(* Logix 5000 project; controller FV vendor 1 type 14 code 217 rev 31.11; software revision 31.00; part 4 of 63 *)

        [1]   // FV12,TEMPERATURE BREAKPOINT A. TIME 1/10 HOURS(ALWAYS=0)
        [15].5   // FV12,Profile Control Flags : This is a conditioning profile
        [29].1   // FV12,Current vessel deferred chilling enabled flag
        [3]   // FV12,TEMPERATURE BREAKPOINT B. TIME 1/10 HOURS(ALWAYS=0)
        [5]   // FV12,TEMPERATURE BREAKPOINT C. TIME 1/10 HOURS(ALWAYS=0)
        [7]   // FV12,TEMPERATURE BREAKPOINT D. TIME 1/10 HOURS(ALWAYS=0)
        [9]   // FV12,TEMPERATURE BREAKPOINT E. TIME 1/10 HOURS(ALWAYS=0)
        [15].9   // FV12,Current vessel deferred chilling manual override
   FV_N123 : INT[50] := ([0] := 13, [2] := 170, [3] := 100, [4] := 190, [5] := 245, [6] := 190, [7] := 275, [8] := 160, [9] := 480, [10] := 160, [11] := 580, [12] := 60, [13] := 32767, [14] := 60, [15] := 64, [17] := -32767, [18] := -32767, [19] := 1680, [22] := 487, [23] := 3, [24] := 5, [25] := 153, [26] := 153, [27] := 487, [30] := 1);   // FV13, CURRENT FV DATA
        [15].2   // FV13,PLC TO FOLLOW RAMP Breakpoints A to B
        [15]   // FV13,FLAGS-PROFILE CONTROL
        [41]   // FV13,Cone ACTUAL TEMPERATURE -DEGREES 'C'*10
        [28]   // FV13,CURRENT VOLUME HL*10
        [15].3   // FV13,PLC TO USE CONE COOLING JACKET
        [24]   // FV13,Phase0=No control 1to6 =Fermenting 8 =Pitching Hold 10 =Maturation 11to16=Conditioning
        [26]   // FV13,Calculated Setpoint 1/10 degrees C
        [30].1   // FV13,Cone Cooling Valve to open
        [30].0   // FV13,Jacket Cooling Valve to open
        [19]   // FV13,Current FV max. fermentation time
        [25]   // FV13,Jacket ACTUAL TEMPERATURE -DEGREES 'C'*10
        [20]   // FV13,Current FV warm conditioning time
        [29]   // FV13,FLAGS - PLC CONTROL
        [10]   // FV13,TEMPERATURE SETPOINT E. 1/10 DEGREE 'C'
        [12]   // FV13,TEMPERATURE SETPOINT F. 1/10 DEGREE 'C'
        [14]   // FV13,TEMPERATURE SETPOINT G. 1/10 DEGREE 'C'
        [30].3   // FV13,Current vessel deferred chilling active
        [0]   // FV13,FV SYSTEM WORKING BUFFER VESSEL NUMBER
        [2]   // FV13,TEMPERATURE SETPOINT A. 1/10 DEGREE 'C'
        [30].4   // FV13,Current vessel final temp.reached
        [4]   // FV13,TEMPERATURE SETPOINT B. 1/10 DEGREE 'C'
        [6]   // FV13,TEMPERATURE SETPOINT C. 1/10 DEGREE 'C'
        [8]   // FV13,TEMPERATURE SETPOINT D. 1/10 DEGREE 'C'
        [22]   // FV13,Current FV total residence time
        [29].0   // FV13,PC TO SAVE TEMPERATURE DATA
        [11]   // FV13,TEMPERATURE BREAKPOINT F. TIME 1/10 HOURS(ALWAYS=0)
        [13]   // FV13,TEMPERATURE BREAKPOINT G. TIME 1/10 HOURS(ALWAYS=0)
        [30].5   // FV13,Current vessel deferred chilling temp.high flag
        [16].1   // FV13,Profile control flag Hold at B.P B
        [16].2   // FV13,Profile control flag Hold at B.P C
        [16].3   // FV13,Profile control flag Hold at B.P D
        [16].4   // FV13,Profile control flag Hold at B.P E
        [16].5   // FV13,Profile control flag Hold at B.P F
        [16].6   // FV13,Profile control flag Hold at B.P G
        [15].4   // FV13,Profile Control Flags : This is a maturation profile
        [27]   // FV13,CURRENT ELAPSED HOURS *10
        [40]   // FV13,FV Routing Status 9=Dirty
        [15].5   // FV13,Profile Control Flags : This is a conditioning profile
        [36]   // FV13,Current vessel time to deferred chlling start (hrs.x10)
        [1]   // FV13,TEMPERATURE BREAKPOINT A. TIME 1/10 HOURS(ALWAYS=0)
        [29].1   // FV13,Current vessel deferred chilling enabled flag
        [3]   // FV13,TEMPERATURE BREAKPOINT B. TIME 1/10 HOURS(ALWAYS=0)
        [5]   // FV13,TEMPERATURE BREAKPOINT C. TIME 1/10 HOURS(ALWAYS=0)
        [7]   // FV13,TEMPERATURE BREAKPOINT D. TIME 1/10 HOURS(ALWAYS=0)
        [9]   // FV13,TEMPERATURE BREAKPOINT E. TIME 1/10 HOURS(ALWAYS=0)
        [15].9   // FV13,Current vessel deferred chilling manual override
   FV_N124 : INT[50] := ([0] := 14, [2] := 170, [3] := 100, [4] := 190, [5] := 258, [6] := 190, [7] := 290, [8] := 160, [9] := 505, [10] := 160, [11] := 605, [12] := 60, [13] := 32767, [14] := 60, [15] := 64, [17] := -32767, [18] := -32767, [19] := 1680, [20] := 8, [22] := 1688, [23] := 3, [24] := 6, [25] := 62, [26] := 60, [27] := 1688, [29] := 2, [30] := 24);   // FV14, CURRENT FV DATA
        [15]   // FV14,FLAGS-PROFILE CONTROL
        [15].2   // FV14,PLC TO FOLLOW RAMP Breakpoints A to B
        [41]   // FV14,Cone ACTUAL TEMPERATURE -DEGREES 'C'*10
        [28]   // FV14,CURRENT VOLUME HL*10
        [30].1   // FV14,Cone Cooling Valve to open
        [15].3   // FV14,PLC TO USE CONE COOLING JACKET
        [24]   // FV14,Phase0=No control 1to6 =Fermenting 8 =Pitching Hold 10 =Maturation 11to16=Conditioning
        [25]   // FV14,Jacket ACTUAL TEMPERATURE -DEGREES 'C'*10
        [26]   // FV14,Calculated Setpoint 1/10 degrees C
        [30].0   // FV14,Jacket Cooling Valve to open
        [19]   // FV14,Current FV max. fermentation time
        [20]   // FV14,Current FV warm conditioning time
        [29]   // FV14,FLAGS - PLC CONTROL
        [0]   // FV14,FV SYSTEM WORKING BUFFER VESSEL NUMBER
        [10]   // FV14,TEMPERATURE SETPOINT E. 1/10 DEGREE 'C'
        [12]   // FV14,TEMPERATURE SETPOINT F. 1/10 DEGREE 'C'
        [2]   // FV14,TEMPERATURE SETPOINT A. 1/10 DEGREE 'C'
        [14]   // FV14,TEMPERATURE SETPOINT G. 1/10 DEGREE 'C'
        [30].3   // FV14,Current vessel deferred chilling active
        [30].4   // FV14,Current vessel final temp.reached
        [4]   // FV14,TEMPERATURE SETPOINT B. 1/10 DEGREE 'C'
        [6]   // FV14,TEMPERATURE SETPOINT C. 1/10 DEGREE 'C'
        [8]   // FV14,TEMPERATURE SETPOINT D. 1/10 DEGREE 'C'
        [22]   // FV14,Current FV total residence time
        [29].0   // FV14,PC TO SAVE TEMPERATURE DATA
        [11]   // FV14,TEMPERATURE BREAKPOINT F. TIME 1/10 HOURS(ALWAYS=0)
        [13]   // FV14,TEMPERATURE BREAKPOINT G. TIME 1/10 HOURS(ALWAYS=0)
        [30].5   // FV14,Current vessel deferred chilling temp.high flag
        [16].1   // FV14,Profile control flag Hold at B.P B
        [16].2   // FV14,Profile control flag Hold at B.P C
        [16].3   // FV14,Profile control flag Hold at B.P D
        [16].4   // FV14,Profile control flag Hold at B.P E
        [16].5   // FV14,Profile control flag Hold at B.P F
        [16].6   // FV14,Profile control flag Hold at B.P G
        [27]   // FV14,CURRENT ELAPSED HOURS *10
        [40]   // FV14,FV Routing Status 9=Dirty
        [15].4   // FV14,Profile Control Flags : This is a maturation profile
        [15].5   // FV14,Profile Control Flags : This is a conditioning profile
        [36]   // FV14,Current vessel time to deferred chlling start (hrs.x10)
        [15].9   // FV14,Current vessel deferred chilling manual override
        [1]   // FV14,TEMPERATURE BREAKPOINT A. TIME 1/10 HOURS(ALWAYS=0)
        [29].1   // FV14,Current vessel deferred chilling enabled flag
        [3]   // FV14,TEMPERATURE BREAKPOINT B. TIME 1/10 HOURS(ALWAYS=0)
        [5]   // FV14,TEMPERATURE BREAKPOINT C. TIME 1/10 HOURS(ALWAYS=0)
        [7]   // FV14,TEMPERATURE BREAKPOINT D. TIME 1/10 HOURS(ALWAYS=0)
        [9]   // FV14,TEMPERATURE BREAKPOINT E. TIME 1/10 HOURS(ALWAYS=0)
   FV_N125 : INT[50] := ([0] := 15, [2] := 170, [3] := 100, [4] := 190, [5] := 270, [6] := 190, [7] := 300, [8] := 160, [9] := 530, [10] := 160, [11] := 630, [12] := 60, [13] := 32767, [14] := 60, [15] := 64, [16] := 20, [17] := -32767, [18] := -32767, [19] := 1680, [22] := 8, [23] := 1, [24] := 1, [25] := 174, [26] := 190, [27] := 8);   // FV15, CURRENT FV DATA
        [15]   // FV15,FLAGS-PROFILE CONTROL
        [15].2   // FV15,PLC TO FOLLOW RAMP Breakpoints A to B
        [41]   // FV15,Cone ACTUAL TEMPERATURE -DEGREES 'C'*10
        [28]   // FV15,CURRENT VOLUME HL*10
        [30].0   // FV15,Jacket Cooling Valve to open
        [30].1   // FV15,Cone Cooling Valve to open
        [15].3   // FV15,PLC TO USE CONE COOLING JACKET
        [24]   // FV15,Phase0=No control 1to6 =Fermenting 8 =Pitching Hold 10 =Maturation 11to16=Conditioning
        [25]   // FV15,Jacket ACTUAL TEMPERATURE -DEGREES 'C'*10
        [26]   // FV15,Calculated Setpoint 1/10 degrees C
        [19]   // FV15,Current FV max. fermentation time
        [20]   // FV15,Current FV warm conditioning time
        [29]   // FV15,FLAGS - PLC CONTROL
        [10]   // FV15,TEMPERATURE SETPOINT E. 1/10 DEGREE 'C'
        [0]   // FV15,FV SYSTEM WORKING BUFFER VESSEL NUMBER
        [2]   // FV15,TEMPERATURE SETPOINT A. 1/10 DEGREE 'C'
        [12]   // FV15,TEMPERATURE SETPOINT F. 1/10 DEGREE 'C'
        [30].4   // FV15,Current vessel final temp.reached
        [14]   // FV15,TEMPERATURE SETPOINT G. 1/10 DEGREE 'C'
        [4]   // FV15,TEMPERATURE SETPOINT B. 1/10 DEGREE 'C'
        [6]   // FV15,TEMPERATURE SETPOINT C. 1/10 DEGREE 'C'
        [8]   // FV15,TEMPERATURE SETPOINT D. 1/10 DEGREE 'C'
        [30].3   // FV15,Current vessel deferred chilling active
        [22]   // FV15,Current FV total residence time
        [29].0   // FV15,PC TO SAVE TEMPERATURE DATA
        [11]   // FV15,TEMPERATURE BREAKPOINT F. TIME 1/10 HOURS(ALWAYS=0)
        [13]   // FV15,TEMPERATURE BREAKPOINT G. TIME 1/10 HOURS(ALWAYS=0)
        [30].5   // FV15,Current vessel deferred chilling temp.high flag
        [16].1   // FV15,Profile control flag Hold at B.P B
        [16].2   // FV15,Profile control flag Hold at B.P C
        [16].3   // FV15,Profile control flag Hold at B.P D
        [16].4   // FV15,Profile control flag Hold at B.P E
        [16].5   // FV15,Profile control flag Hold at B.P F
        [16].6   // FV15,Profile control flag Hold at B.P G
        [15].4   // FV15,Profile Control Flags : This is a maturation profile
        [15].5   // FV15,Profile Control Flags : This is a conditioning profile
        [27]   // FV15,CURRENT ELAPSED HOURS *10
        [40]   // FV15,FV Routing Status 9=Dirty
        [36]   // FV15,Current vessel time to deferred chlling start (hrs.x10)
        [15].9   // FV15,Current vessel deferred chilling manual override
        [1]   // FV15,TEMPERATURE BREAKPOINT A. TIME 1/10 HOURS(ALWAYS=0)
        [29].1   // FV15,Current vessel deferred chilling enabled flag
        [3]   // FV15,TEMPERATURE BREAKPOINT B. TIME 1/10 HOURS(ALWAYS=0)
        [5]   // FV15,TEMPERATURE BREAKPOINT C. TIME 1/10 HOURS(ALWAYS=0)
        [7]   // FV15,TEMPERATURE BREAKPOINT D. TIME 1/10 HOURS(ALWAYS=0)
        [9]   // FV15,TEMPERATURE BREAKPOINT E. TIME 1/10 HOURS(ALWAYS=0)
   FV_N126 : INT[50] := ([0] := 16, [1] := -32767, [2] := -32767, [3] := -32767, [4] := -32767, [5] := -32767, [6] := -32767, [7] := -32767, [8] := -32767, [9] := -32767, [10] := -32767, [11] := -32767, [12] := -32767, [13] := -32767, [14] := -32767, [15] := -32767, [16] := -32767, [17] := -32767, [18] := -32767, [19] := -32767, [20] := -32767, [21] := -32767, [22] := -32767, [23] := 2, [25] := 201, [30] := 32);   // FV16, CURRENT FV DATA
        [15]   // FV16,FLAGS-PROFILE CONTROL
        [15].2   // FV16,PLC TO FOLLOW RAMP Breakpoints A to B
        [41]   // FV16,Cone ACTUAL TEMPERATURE -DEGREES 'C'*10
        [28]   // FV16,CURRENT VOLUME HL*10
        [25]   // FV16,Jacket ACTUAL TEMPERATURE -DEGREES 'C'*10
        [15].3   // FV16,PLC TO USE CONE COOLING JACKET
        [30].0   // FV16,Jacket Cooling Valve to open
        [26]   // FV16,Calculated Setpoint 1/10 degrees C
        [30].1   // FV16,Cone Cooling Valve to open
        [24]   // FV16,Phase0=No control 1to6 =Fermenting 8 =Pitching Hold 10 =Maturation 11to16=Conditioning
        [19]   // FV16,Current FV max. fermentation time
        [20]   // FV16,Current FV warm conditioning time
        [29]   // FV16,FLAGS - PLC CONTROL
        [10]   // FV16,TEMPERATURE SETPOINT E. 1/10 DEGREE 'C'
        [12]   // FV16,TEMPERATURE SETPOINT F. 1/10 DEGREE 'C'
        [14]   // FV16,TEMPERATURE SETPOINT G. 1/10 DEGREE 'C'
        [0]   // FV16,FV SYSTEM WORKING BUFFER VESSEL NUMBER
        [2]   // FV16,TEMPERATURE SETPOINT A. 1/10 DEGREE 'C'
        [30].4   // FV16,Current vessel final temp.reached
        [4]   // FV16,TEMPERATURE SETPOINT B. 1/10 DEGREE 'C'
        [6]   // FV16,TEMPERATURE SETPOINT C. 1/10 DEGREE 'C'
        [8]   // FV16,TEMPERATURE SETPOINT D. 1/10 DEGREE 'C'
        [30].3   // FV16,Current vessel deferred chilling active
        [22]   // FV16,Current FV total residence time
        [29].0   // FV16,PC TO SAVE TEMPERATURE DATA
        [11]   // FV16,TEMPERATURE BREAKPOINT F. TIME 1/10 HOURS(ALWAYS=0)
        [13]   // FV16,TEMPERATURE BREAKPOINT G. TIME 1/10 HOURS(ALWAYS=0)
        [30].5   // FV16,Current vessel deferred chilling temp.high flag
        [36]   // FV16,Current vessel time to deferred chlling start (hrs.x10)
        [15].4   // FV16,Profile Control Flags : This is a maturation profile
        [15].5   // FV16,Profile Control Flags : This is a conditioning profile
        [16].1   // FV16,Profile control flag Hold at B.P B
        [16].2   // FV16,Profile control flag Hold at B.P C
        [16].3   // FV16,Profile control flag Hold at B.P D
        [16].4   // FV16,Profile control flag Hold at B.P E
        [16].5   // FV16,Profile control flag Hold at B.P F
        [16].6   // FV16,Profile control flag Hold at B.P G
        [27]   // FV16,CURRENT ELAPSED HOURS *10
        [40]   // FV16,FV Routing Status 9=Dirty
        [15].9   // FV16,Current vessel deferred chilling manual override
        [1]   // FV16,TEMPERATURE BREAKPOINT A. TIME 1/10 HOURS(ALWAYS=0)
        [29].1   // FV16,Current vessel deferred chilling enabled flag
        [3]   // FV16,TEMPERATURE BREAKPOINT B. TIME 1/10 HOURS(ALWAYS=0)
        [5]   // FV16,TEMPERATURE BREAKPOINT C. TIME 1/10 HOURS(ALWAYS=0)
        [7]   // FV16,TEMPERATURE BREAKPOINT D. TIME 1/10 HOURS(ALWAYS=0)
        [9]   // FV16,TEMPERATURE BREAKPOINT E. TIME 1/10 HOURS(ALWAYS=0)
   FV_N127 : INT[50] := ([0] := 17, [1] := -32767, [2] := -32767, [3] := -32767, [4] := -32767, [5] := -32767, [6] := -32767, [7] := -32767, [8] := -32767, [9] := -32767, [10] := -32767, [11] := -32767, [12] := -32767, [13] := -32767, [14] := -32767, [15] := -32767, [16] := -32767, [17] := -32767, [18] := -32767, [19] := -32767, [20] := -32767, [21] := -32767, [22] := -32767, [23] := 2, [25] := 203, [30] := 32);   // FV17, CURRENT FV DATA
        [15]   // FV17,FLAGS-PROFILE CONTROL
        [15].2   // FV17,PLC TO FOLLOW RAMP Breakpoints A to B
        [41]   // FV17,Cone ACTUAL TEMPERATURE -DEGREES 'C'*10
        [25]   // FV17,Jacket ACTUAL TEMPERATURE -DEGREES 'C'*10
        [28]   // FV17,CURRENT VOLUME HL*10
        [15].3   // FV17,PLC TO USE CONE COOLING JACKET
        [30].0   // FV17,Jacket Cooling Valve to open
        [26]   // FV17,Calculated Setpoint 1/10 degrees C
        [24]   // FV17,Phase0=No control 1to6 =Fermenting 8 =Pitching Hold 10 =Maturation 11to16=Conditioning
        [30].1   // FV17,Cone Cooling Valve to open
        [19]   // FV17,Current FV max. fermentation time
        [10]   // FV17,TEMPERATURE SETPOINT E. 1/10 DEGREE 'C'
        [20]   // FV17,Current FV warm conditioning time
        [12]   // FV17,TEMPERATURE SETPOINT F. 1/10 DEGREE 'C'
        [29]   // FV17,FLAGS - PLC CONTROL
        [14]   // FV17,TEMPERATURE SETPOINT G. 1/10 DEGREE 'C'
        [0]   // FV17,FV SYSTEM WORKING BUFFER VESSEL NUMBER
        [2]   // FV17,TEMPERATURE SETPOINT A. 1/10 DEGREE 'C'
        [30].4   // FV17,Current vessel final temp.reached
        [4]   // FV17,TEMPERATURE SETPOINT B. 1/10 DEGREE 'C'
        [6]   // FV17,TEMPERATURE SETPOINT C. 1/10 DEGREE 'C'
        [8]   // FV17,TEMPERATURE SETPOINT D. 1/10 DEGREE 'C'
        [30].3   // FV17,Current vessel deferred chilling active
        [22]   // FV17,Current FV total residence time
        [29].0   // FV17,PC TO SAVE TEMPERATURE DATA
        [36]   // FV17,Current vessel time to deferred chlling start (hrs.x10)
        [11]   // FV17,TEMPERATURE BREAKPOINT F. TIME 1/10 HOURS(ALWAYS=0)
        [13]   // FV17,TEMPERATURE BREAKPOINT G. TIME 1/10 HOURS(ALWAYS=0)
        [30].5   // FV17,Current vessel deferred chilling temp.high flag
        [15].4   // FV17,Profile Control Flags : This is a maturation profile
        [27]   // FV17,CURRENT ELAPSED HOURS *10
        [40]   // FV17,FV Routing Status 9=Dirty
        [16].1   // FV17,Profile control flag Hold at B.P B
        [15].5   // FV17,Profile Control Flags : This is a conditioning profile
        [16].2   // FV17,Profile control flag Hold at B.P C
        [16].3   // FV17,Profile control flag Hold at B.P D
        [16].4   // FV17,Profile control flag Hold at B.P E
        [16].5   // FV17,Profile control flag Hold at B.P F
        [16].6   // FV17,Profile control flag Hold at B.P G
        [15].9   // FV17,Current vessel deferred chilling manual override
        [1]   // FV17,TEMPERATURE BREAKPOINT A. TIME 1/10 HOURS(ALWAYS=0)
        [29].1   // FV17,Current vessel deferred chilling enabled flag
        [3]   // FV17,TEMPERATURE BREAKPOINT B. TIME 1/10 HOURS(ALWAYS=0)
        [5]   // FV17,TEMPERATURE BREAKPOINT C. TIME 1/10 HOURS(ALWAYS=0)
        [7]   // FV17,TEMPERATURE BREAKPOINT D. TIME 1/10 HOURS(ALWAYS=0)
        [9]   // FV17,TEMPERATURE BREAKPOINT E. TIME 1/10 HOURS(ALWAYS=0)
   FV_N128 : INT[50] := ([0] := 18, [1] := -32767, [2] := -32767, [3] := -32767, [4] := -32767, [5] := -32767, [6] := -32767, [7] := -32767, [8] := -32767, [9] := -32767, [10] := -32767, [11] := -32767, [12] := -32767, [13] := -32767, [14] := -32767, [15] := -32767, [16] := -32767, [17] := -32767, [18] := -32767, [19] := -32767, [20] := -32767, [21] := -32767, [22] := -32767, [23] := 2, [25] := 216, [30] := 32);   // FV18, CURRENT FV DATA
        [15]   // FV18,FLAGS-PROFILE CONTROL
        [15].2   // FV18,PLC TO FOLLOW RAMP Breakpoints A to B
        [25]   // FV18,Jacket ACTUAL TEMPERATURE -DEGREES 'C'*10
        [41]   // FV18,Cone ACTUAL TEMPERATURE -DEGREES 'C'*10
        [28]   // FV18,CURRENT VOLUME HL*10
        [15].3   // FV18,PLC TO USE CONE COOLING JACKET
        [26]   // FV18,Calculated Setpoint 1/10 degrees C
        [30].0   // FV18,Jacket Cooling Valve to open
        [30].1   // FV18,Cone Cooling Valve to open
        [24]   // FV18,Phase0=No control 1to6 =Fermenting 8 =Pitching Hold 10 =Maturation 11to16=Conditioning
        [19]   // FV18,Current FV max. fermentation time
        [20]   // FV18,Current FV warm conditioning time
        [10]   // FV18,TEMPERATURE SETPOINT E. 1/10 DEGREE 'C'
        [12]   // FV18,TEMPERATURE SETPOINT F. 1/10 DEGREE 'C'
        [14]   // FV18,TEMPERATURE SETPOINT G. 1/10 DEGREE 'C'
        [29]   // FV18,FLAGS - PLC CONTROL
        [0]   // FV18,FV SYSTEM WORKING BUFFER VESSEL NUMBER
        [2]   // FV18,TEMPERATURE SETPOINT A. 1/10 DEGREE 'C'
        [30].4   // FV18,Current vessel final temp.reached
        [4]   // FV18,TEMPERATURE SETPOINT B. 1/10 DEGREE 'C'
        [6]   // FV18,TEMPERATURE SETPOINT C. 1/10 DEGREE 'C'
        [8]   // FV18,TEMPERATURE SETPOINT D. 1/10 DEGREE 'C'
        [30].3   // FV18,Current vessel deferred chilling active
        [22]   // FV18,Current FV total residence time
        [29].0   // FV18,PC TO SAVE TEMPERATURE DATA
        [36]   // FV18,Current vessel time to deferred chlling start (hrs.x10)
        [15].4   // FV18,Profile Control Flags : This is a maturation profile
        [15].5   // FV18,Profile Control Flags : This is a conditioning profile
        [11]   // FV18,TEMPERATURE BREAKPOINT F. TIME 1/10 HOURS(ALWAYS=0)
        [13]   // FV18,TEMPERATURE BREAKPOINT G. TIME 1/10 HOURS(ALWAYS=0)
        [30].5   // FV18,Current vessel deferred chilling temp.high flag
        [16].1   // FV18,Profile control flag Hold at B.P B
        [16].2   // FV18,Profile control flag Hold at B.P C
        [16].3   // FV18,Profile control flag Hold at B.P D
        [16].4   // FV18,Profile control flag Hold at B.P E
        [27]   // FV18,CURRENT ELAPSED HOURS *10
        [16].5   // FV18,Profile control flag Hold at B.P F
        [40]   // FV18,FV Routing Status 9=Dirty
        [16].6   // FV18,Profile control flag Hold at B.P G
        [15].9   // FV18,Current vessel deferred chilling manual override
        [1]   // FV18,TEMPERATURE BREAKPOINT A. TIME 1/10 HOURS(ALWAYS=0)
        [29].1   // FV18,Current vessel deferred chilling enabled flag
        [3]   // FV18,TEMPERATURE BREAKPOINT B. TIME 1/10 HOURS(ALWAYS=0)
        [5]   // FV18,TEMPERATURE BREAKPOINT C. TIME 1/10 HOURS(ALWAYS=0)
        [7]   // FV18,TEMPERATURE BREAKPOINT D. TIME 1/10 HOURS(ALWAYS=0)
        [9]   // FV18,TEMPERATURE BREAKPOINT E. TIME 1/10 HOURS(ALWAYS=0)
   FV_N129 : INT[50] := ([0] := 19, [1] := -32767, [2] := -32767, [3] := -32767, [4] := -32767, [5] := -32767, [6] := -32767, [7] := -32767, [8] := -32767, [9] := -32767, [10] := -32767, [11] := -32767, [12] := -32767, [13] := -32767, [14] := -32767, [15] := -32767, [16] := -32767, [17] := -32767, [18] := -32767, [19] := -32767, [20] := -32767, [21] := -32767, [22] := -32767, [23] := 2, [25] := 219, [30] := 32);   // FV19, CURRENT FV DATA
        [15]   // FV19,FLAGS-PROFILE CONTROL
        [15].2   // FV19,PLC TO FOLLOW RAMP Breakpoints A to B
        [25]   // FV19,Jacket ACTUAL TEMPERATURE -DEGREES 'C'*10
        [41]   // FV19,Cone ACTUAL TEMPERATURE -DEGREES 'C'*10
        [28]   // FV19,CURRENT VOLUME HL*10
        [30].1   // FV19,Cone Cooling Valve to open
        [15].3   // FV19,PLC TO USE CONE COOLING JACKET
        [26]   // FV19,Calculated Setpoint 1/10 degrees C
        [30].0   // FV19,Jacket Cooling Valve to open
        [15].5   // FV19,Profile Control Flags : This is a conditioning profile
        [24]   // FV19,Phase0=No control 1to6 =Fermenting 8 =Pitching Hold 10 =Maturation 11to16=Conditioning
        [10]   // FV19,TEMPERATURE SETPOINT E. 1/10 DEGREE 'C'
        [19]   // FV19,Current FV max. fermentation time
        [20]   // FV19,Current FV warm conditioning time
        [12]   // FV19,TEMPERATURE SETPOINT F. 1/10 DEGREE 'C'
        [14]   // FV19,TEMPERATURE SETPOINT G. 1/10 DEGREE 'C'
        [29]   // FV19,FLAGS - PLC CONTROL
        [0]   // FV19,FV SYSTEM WORKING BUFFER VESSEL NUMBER
        [2]   // FV19,TEMPERATURE SETPOINT A. 1/10 DEGREE 'C'
        [30].4   // FV19,Current vessel final temp.reached
        [30].3   // FV19,Current vessel deferred chilling active
        [4]   // FV19,TEMPERATURE SETPOINT B. 1/10 DEGREE 'C'
        [6]   // FV19,TEMPERATURE SETPOINT C. 1/10 DEGREE 'C'
        [8]   // FV19,TEMPERATURE SETPOINT D. 1/10 DEGREE 'C'
        [15].4   // FV19,Profile Control Flags : This is a maturation profile
        [22]   // FV19,Current FV total residence time
        [29].0   // FV19,PC TO SAVE TEMPERATURE DATA
        [36]   // FV19,Current vessel time to deferred chlling start (hrs.x10)
        [11]   // FV19,TEMPERATURE BREAKPOINT F. TIME 1/10 HOURS(ALWAYS=0)
        [13]   // FV19,TEMPERATURE BREAKPOINT G. TIME 1/10 HOURS(ALWAYS=0)
        [30].5   // FV19,Current vessel deferred chilling temp.high flag
        [27]   // FV19,CURRENT ELAPSED HOURS *10
        [16].1   // FV19,Profile control flag Hold at B.P B
        [16].2   // FV19,Profile control flag Hold at B.P C
        [16].3   // FV19,Profile control flag Hold at B.P D
        [16].4   // FV19,Profile control flag Hold at B.P E
        [16].5   // FV19,Profile control flag Hold at B.P F
        [16].6   // FV19,Profile control flag Hold at B.P G
        [40]   // FV19,FV Routing Status 9=Dirty
        [15].9   // FV19,Current vessel deferred chilling manual override
        [1]   // FV19,TEMPERATURE BREAKPOINT A. TIME 1/10 HOURS(ALWAYS=0)
        [29].1   // FV19,Current vessel deferred chilling enabled flag
        [3]   // FV19,TEMPERATURE BREAKPOINT B. TIME 1/10 HOURS(ALWAYS=0)
        [5]   // FV19,TEMPERATURE BREAKPOINT C. TIME 1/10 HOURS(ALWAYS=0)
        [7]   // FV19,TEMPERATURE BREAKPOINT D. TIME 1/10 HOURS(ALWAYS=0)
        [9]   // FV19,TEMPERATURE BREAKPOINT E. TIME 1/10 HOURS(ALWAYS=0)
   FV_N13 : INT[255] := ([3] := 6, [16] := 123, [19] := 17);   // PLC>ME Inter PLC comms traf fic inbound
        [2].0   // MVSYSTEM>Me Acknowledgement of request to set MV status to ageing
        [18].0   // CTSYSTEM>Me Acknowledgement of request to set CT status to ageing
        [19]   // CTSYSTEM>Me Number of cooling valves open in CT system
        [3]   // MVSYSTEM>Me Number of cooling valves open in MV system
        [2]   // MVSYSTEM>Me Request acknowledgement flags
   FV_N130 : INT[50] := ([0] := 20, [1] := -32767, [2] := -32767, [3] := -32767, [4] := -32767, [5] := -32767, [6] := -32767, [7] := -32767, [8] := -32767, [9] := -32767, [10] := -32767, [11] := -32767, [12] := -32767, [13] := -32767, [14] := -32767, [15] := -32767, [16] := -32767, [17] := -32767, [18] := -32767, [19] := -32767, [20] := -32767, [21] := -32767, [22] := -32767, [23] := 2, [25] := 218, [30] := 32);   // FV20, CURRENT FV DATA
        [15]   // FV20,FLAGS-PROFILE CONTROL
        [15].2   // FV20,PLC TO FOLLOW RAMP Breakpoints A to B
        [25]   // FV20,Jacket ACTUAL TEMPERATURE -DEGREES 'C'*10
        [41]   // FV20,Cone ACTUAL TEMPERATURE -DEGREES 'C'*10
        [28]   // FV20,CURRENT VOLUME HL*10
        [30].1   // FV20,Cone Cooling Valve to open
        [15].3   // FV20,PLC TO USE CONE COOLING JACKET
        [26]   // FV20,Calculated Setpoint 1/10 degrees C
        [15].5   // FV20,Profile Control Flags : This is a conditioning profile
        [30].0   // FV20,Jacket Cooling Valve to open
        [24]   // FV20,Phase0=No control 1to6 =Fermenting 8 =Pitching Hold 10 =Maturation 11to16=Conditioning
        [19]   // FV20,Current FV max. fermentation time
        [10]   // FV20,TEMPERATURE SETPOINT E. 1/10 DEGREE 'C'
        [12]   // FV20,TEMPERATURE SETPOINT F. 1/10 DEGREE 'C'
        [14]   // FV20,TEMPERATURE SETPOINT G. 1/10 DEGREE 'C'
        [15].4   // FV20,Profile Control Flags : This is a maturation profile
        [20]   // FV20,Current FV warm conditioning time
        [30].3   // FV20,Current vessel deferred chilling active
        [0]   // FV20,FV SYSTEM WORKING BUFFER VESSEL NUMBER
        [29]   // FV20,FLAGS - PLC CONTROL
        [2]   // FV20,TEMPERATURE SETPOINT A. 1/10 DEGREE 'C'
        [30].4   // FV20,Current vessel final temp.reached
        [4]   // FV20,TEMPERATURE SETPOINT B. 1/10 DEGREE 'C'
        [6]   // FV20,TEMPERATURE SETPOINT C. 1/10 DEGREE 'C'
        [8]   // FV20,TEMPERATURE SETPOINT D. 1/10 DEGREE 'C'
        [36]   // FV20,Current vessel time to deferred chlling start (hrs.x10)
        [22]   // FV20,Current FV total residence time
        [29].0   // FV20,PC TO SAVE TEMPERATURE DATA
        [27]   // FV20,CURRENT ELAPSED HOURS *10
        [40]   // FV20,FV Routing Status 9=Dirty
        [11]   // FV20,TEMPERATURE BREAKPOINT F. TIME 1/10 HOURS(ALWAYS=0)
        [13]   // FV20,TEMPERATURE BREAKPOINT G. TIME 1/10 HOURS(ALWAYS=0)
        [30].5   // FV20,Current vessel deferred chilling temp.high flag
        [16].1   // FV20,Profile control flag Hold at B.P B
        [16].2   // FV20,Profile control flag Hold at B.P C
        [16].3   // FV20,Profile control flag Hold at B.P D
        [16].4   // FV20,Profile control flag Hold at B.P E
        [16].5   // FV20,Profile control flag Hold at B.P F
        [16].6   // FV20,Profile control flag Hold at B.P G
        [15].9   // FV20,Current vessel deferred chilling manual override
        [1]   // FV20,TEMPERATURE BREAKPOINT A. TIME 1/10 HOURS(ALWAYS=0)
        [29].1   // FV20,Current vessel deferred chilling enabled flag
        [3]   // FV20,TEMPERATURE BREAKPOINT B. TIME 1/10 HOURS(ALWAYS=0)
        [5]   // FV20,TEMPERATURE BREAKPOINT C. TIME 1/10 HOURS(ALWAYS=0)
        [7]   // FV20,TEMPERATURE BREAKPOINT D. TIME 1/10 HOURS(ALWAYS=0)
        [9]   // FV20,TEMPERATURE BREAKPOINT E. TIME 1/10 HOURS(ALWAYS=0)
   FV_N131 : INT[50] := ([0] := 21, [1] := -32767, [2] := -32767, [3] := -32767, [4] := -32767, [5] := -32767, [6] := -32767, [7] := -32767, [8] := -32767, [9] := -32767, [10] := -32767, [11] := -32767, [12] := -32767, [13] := -32767, [14] := -32767, [15] := -32767, [16] := -32767, [17] := -32767, [18] := -32767, [19] := -32767, [20] := -32767, [21] := -32767, [22] := -32767, [23] := 2, [25] := 221, [30] := 32);   // FV21, CURRENT FV DATA
        [15]   // FV21,FLAGS-PROFILE CONTROL
        [15].5   // FV21,Profile Control Flags : This is a conditioning profile
        [25]   // FV21,Jacket ACTUAL TEMPERATURE -DEGREES 'C'*10
        [15].2   // FV21,PLC TO FOLLOW RAMP Breakpoints A to B
        [41]   // FV21,Cone ACTUAL TEMPERATURE -DEGREES 'C'*10
        [28]   // FV21,CURRENT VOLUME HL*10
        [15].3   // FV21,PLC TO USE CONE COOLING JACKET
        [30].1   // FV21,Cone Cooling Valve to open
        [26]   // FV21,Calculated Setpoint 1/10 degrees C
        [19]   // FV21,Current FV max. fermentation time
        [20]   // FV21,Current FV warm conditioning time
        [30].0   // FV21,Jacket Cooling Valve to open
        [24]   // FV21,Phase0=No control 1to6 =Fermenting 8 =Pitching Hold 10 =Maturation 11to16=Conditioning
        [15].4   // FV21,Profile Control Flags : This is a maturation profile
        [10]   // FV21,TEMPERATURE SETPOINT E. 1/10 DEGREE 'C'
        [12]   // FV21,TEMPERATURE SETPOINT F. 1/10 DEGREE 'C'
        [14]   // FV21,TEMPERATURE SETPOINT G. 1/10 DEGREE 'C'
        [30].3   // FV21,Current vessel deferred chilling active
        [0]   // FV21,FV SYSTEM WORKING BUFFER VESSEL NUMBER
        [2]   // FV21,TEMPERATURE SETPOINT A. 1/10 DEGREE 'C'
        [30].4   // FV21,Current vessel final temp.reached
        [4]   // FV21,TEMPERATURE SETPOINT B. 1/10 DEGREE 'C'
        [6]   // FV21,TEMPERATURE SETPOINT C. 1/10 DEGREE 'C'
        [8]   // FV21,TEMPERATURE SETPOINT D. 1/10 DEGREE 'C'
        [29]   // FV21,FLAGS - PLC CONTROL
        [36]   // FV21,Current vessel time to deferred chlling start (hrs.x10)
        [22]   // FV21,Current FV total residence time
        [27]   // FV21,CURRENT ELAPSED HOURS *10
        [29].0   // FV21,PC TO SAVE TEMPERATURE DATA
        [40]   // FV21,FV Routing Status 9=Dirty
        [16].1   // FV21,Profile control flag Hold at B.P B
        [16].2   // FV21,Profile control flag Hold at B.P C
        [11]   // FV21,TEMPERATURE BREAKPOINT F. TIME 1/10 HOURS(ALWAYS=0)
        [16].3   // FV21,Profile control flag Hold at B.P D
        [16].4   // FV21,Profile control flag Hold at B.P E
        [13]   // FV21,TEMPERATURE BREAKPOINT G. TIME 1/10 HOURS(ALWAYS=0)
        [30].5   // FV21,Current vessel deferred chilling temp.high flag
        [16].5   // FV21,Profile control flag Hold at B.P F
        [16].6   // FV21,Profile control flag Hold at B.P G
        [15].9   // FV21,Current vessel deferred chilling manual override
        [1]   // FV21,TEMPERATURE BREAKPOINT A. TIME 1/10 HOURS(ALWAYS=0)
        [29].1   // FV21,Current vessel deferred chilling enabled flag
        [3]   // FV21,TEMPERATURE BREAKPOINT B. TIME 1/10 HOURS(ALWAYS=0)
        [5]   // FV21,TEMPERATURE BREAKPOINT C. TIME 1/10 HOURS(ALWAYS=0)
        [7]   // FV21,TEMPERATURE BREAKPOINT D. TIME 1/10 HOURS(ALWAYS=0)
        [9]   // FV21,TEMPERATURE BREAKPOINT E. TIME 1/10 HOURS(ALWAYS=0)
   FV_N132 : INT[50] := ([0] := 22, [1] := -32767, [2] := -32767, [3] := -32767, [4] := -32767, [5] := -32767, [6] := -32767, [7] := -32767, [8] := -32767, [9] := -32767, [10] := -32767, [11] := -32767, [12] := -32767, [13] := -32767, [14] := -32767, [15] := -32767, [16] := -32767, [17] := -32767, [18] := -32767, [19] := -32767, [20] := -32767, [21] := -32767, [22] := -32767, [23] := 2, [25] := 164, [30] := 32);   // FV22, CURRENT FV DATA
        [15]   // FV22,FLAGS-PROFILE CONTROL
        [15].5   // FV22,Profile Control Flags : This is a conditioning profile
        [25]   // FV22,Jacket ACTUAL TEMPERATURE -DEGREES 'C'*10
        [15].2   // FV22,PLC TO FOLLOW RAMP Breakpoints A to B
        [41]   // FV22,Cone ACTUAL TEMPERATURE -DEGREES 'C'*10
        [28]   // FV22,CURRENT VOLUME HL*10
        [19]   // FV22,Current FV max. fermentation time
        [15].3   // FV22,PLC TO USE CONE COOLING JACKET
        [30].1   // FV22,Cone Cooling Valve to open
        [20]   // FV22,Current FV warm conditioning time
        [26]   // FV22,Calculated Setpoint 1/10 degrees C
        [30].0   // FV22,Jacket Cooling Valve to open
        [30].3   // FV22,Current vessel deferred chilling active
        [10]   // FV22,TEMPERATURE SETPOINT E. 1/10 DEGREE 'C'
        [24]   // FV22,Phase0=No control 1to6 =Fermenting 8 =Pitching Hold 10 =Maturation 11to16=Conditioning
        [12]   // FV22,TEMPERATURE SETPOINT F. 1/10 DEGREE 'C'
        [14]   // FV22,TEMPERATURE SETPOINT G. 1/10 DEGREE 'C'
        [15].4   // FV22,Profile Control Flags : This is a maturation profile
        [36]   // FV22,Current vessel time to deferred chlling start (hrs.x10)
        [0]   // FV22,FV SYSTEM WORKING BUFFER VESSEL NUMBER
        [2]   // FV22,TEMPERATURE SETPOINT A. 1/10 DEGREE 'C'
        [30].4   // FV22,Current vessel final temp.reached
        [4]   // FV22,TEMPERATURE SETPOINT B. 1/10 DEGREE 'C'
        [6]   // FV22,TEMPERATURE SETPOINT C. 1/10 DEGREE 'C'
        [8]   // FV22,TEMPERATURE SETPOINT D. 1/10 DEGREE 'C'
        [29]   // FV22,FLAGS - PLC CONTROL
        [27]   // FV22,CURRENT ELAPSED HOURS *10
        [40]   // FV22,FV Routing Status 9=Dirty
        [22]   // FV22,Current FV total residence time
        [16].1   // FV22,Profile control flag Hold at B.P B
        [29].0   // FV22,PC TO SAVE TEMPERATURE DATA
        [16].2   // FV22,Profile control flag Hold at B.P C
        [16].3   // FV22,Profile control flag Hold at B.P D
        [16].4   // FV22,Profile control flag Hold at B.P E
        [16].5   // FV22,Profile control flag Hold at B.P F
        [16].6   // FV22,Profile control flag Hold at B.P G
        [11]   // FV22,TEMPERATURE BREAKPOINT F. TIME 1/10 HOURS(ALWAYS=0)
        [13]   // FV22,TEMPERATURE BREAKPOINT G. TIME 1/10 HOURS(ALWAYS=0)
        [30].5   // FV22,Current vessel deferred chilling temp.high flag
        [15].9   // FV22,Current vessel deferred chilling manual override
        [1]   // FV22,TEMPERATURE BREAKPOINT A. TIME 1/10 HOURS(ALWAYS=0)
        [29].1   // FV22,Current vessel deferred chilling enabled flag
        [3]   // FV22,TEMPERATURE BREAKPOINT B. TIME 1/10 HOURS(ALWAYS=0)
        [5]   // FV22,TEMPERATURE BREAKPOINT C. TIME 1/10 HOURS(ALWAYS=0)
        [7]   // FV22,TEMPERATURE BREAKPOINT D. TIME 1/10 HOURS(ALWAYS=0)
        [9]   // FV22,TEMPERATURE BREAKPOINT E. TIME 1/10 HOURS(ALWAYS=0)
   FV_N133 : INT[50] := ([0] := 23, [1] := -32767, [2] := -32767, [3] := -32767, [4] := -32767, [5] := -32767, [6] := -32767, [7] := -32767, [8] := -32767, [9] := -32767, [10] := -32767, [11] := -32767, [12] := -32767, [13] := -32767, [14] := -32767, [15] := -32767, [16] := -32767, [17] := -32767, [18] := -32767, [19] := -32767, [20] := -32767, [21] := -32767, [22] := -32767, [23] := 2, [25] := 212, [30] := 32);   // FV23, CURRENT FV DATA
        [15]   // FV23,FLAGS-PROFILE CONTROL
        [15].5   // FV23,Profile Control Flags : This is a conditioning profile
        [25]   // FV23,Jacket ACTUAL TEMPERATURE -DEGREES 'C'*10
        [15].2   // FV23,PLC TO FOLLOW RAMP Breakpoints A to B
        [41]   // FV23,Cone ACTUAL TEMPERATURE -DEGREES 'C'*10
        [30].3   // FV23,Current vessel deferred chilling active
        [28]   // FV23,CURRENT VOLUME HL*10
        [15].4   // FV23,Profile Control Flags : This is a maturation profile
        [30].1   // FV23,Cone Cooling Valve to open
        [19]   // FV23,Current FV max. fermentation time
        [15].3   // FV23,PLC TO USE CONE COOLING JACKET
        [20]   // FV23,Current FV warm conditioning time
        [26]   // FV23,Calculated Setpoint 1/10 degrees C
        [30].0   // FV23,Jacket Cooling Valve to open
        [10]   // FV23,TEMPERATURE SETPOINT E. 1/10 DEGREE 'C'
        [12]   // FV23,TEMPERATURE SETPOINT F. 1/10 DEGREE 'C'
        [24]   // FV23,Phase0=No control 1to6 =Fermenting 8 =Pitching Hold 10 =Maturation 11to16=Conditioning
        [14]   // FV23,TEMPERATURE SETPOINT G. 1/10 DEGREE 'C'
        [0]   // FV23,FV SYSTEM WORKING BUFFER VESSEL NUMBER
        [36]   // FV23,Current vessel time to deferred chlling start (hrs.x10)
        [2]   // FV23,TEMPERATURE SETPOINT A. 1/10 DEGREE 'C'
        [30].4   // FV23,Current vessel final temp.reached
        [4]   // FV23,TEMPERATURE SETPOINT B. 1/10 DEGREE 'C'
        [6]   // FV23,TEMPERATURE SETPOINT C. 1/10 DEGREE 'C'
        [8]   // FV23,TEMPERATURE SETPOINT D. 1/10 DEGREE 'C'
        [29]   // FV23,FLAGS - PLC CONTROL
        [27]   // FV23,CURRENT ELAPSED HOURS *10
        [40]   // FV23,FV Routing Status 9=Dirty
        [22]   // FV23,Current FV total residence time
        [29].0   // FV23,PC TO SAVE TEMPERATURE DATA
        [16].1   // FV23,Profile control flag Hold at B.P B
        [16].2   // FV23,Profile control flag Hold at B.P C
        [16].3   // FV23,Profile control flag Hold at B.P D
        [16].4   // FV23,Profile control flag Hold at B.P E
        [16].5   // FV23,Profile control flag Hold at B.P F
        [16].6   // FV23,Profile control flag Hold at B.P G
        [11]   // FV23,TEMPERATURE BREAKPOINT F. TIME 1/10 HOURS(ALWAYS=0)
        [13]   // FV23,TEMPERATURE BREAKPOINT G. TIME 1/10 HOURS(ALWAYS=0)
        [30].5   // FV23,Current vessel deferred chilling temp.high flag
        [15].9   // FV23,Current vessel deferred chilling manual override
        [1]   // FV23,TEMPERATURE BREAKPOINT A. TIME 1/10 HOURS(ALWAYS=0)
        [29].1   // FV23,Current vessel deferred chilling enabled flag
        [3]   // FV23,TEMPERATURE BREAKPOINT B. TIME 1/10 HOURS(ALWAYS=0)
        [5]   // FV23,TEMPERATURE BREAKPOINT C. TIME 1/10 HOURS(ALWAYS=0)
        [7]   // FV23,TEMPERATURE BREAKPOINT D. TIME 1/10 HOURS(ALWAYS=0)
        [9]   // FV23,TEMPERATURE BREAKPOINT E. TIME 1/10 HOURS(ALWAYS=0)
   FV_N134 : INT[50] := ([0] := 24, [1] := -32767, [2] := -32767, [3] := -32767, [4] := -32767, [5] := -32767, [6] := -32767, [7] := -32767, [8] := -32767, [9] := -32767, [10] := -32767, [11] := -32767, [12] := -32767, [13] := -32767, [14] := -32767, [15] := -32767, [16] := -32767, [17] := -32767, [18] := -32767, [19] := -32767, [20] := -32767, [21] := -32767, [22] := -32767, [23] := 2, [25] := 216, [30] := 32);   // FV24, CURRENT FV DATA
        [15]   // FV24,FLAGS-PROFILE CONTROL
        [15].4   // FV24,Profile Control Flags : This is a maturation profile
        [25]   // FV24,Jacket ACTUAL TEMPERATURE -DEGREES 'C'*10
        [15].5   // FV24,Profile Control Flags : This is a conditioning profile
        [15].2   // FV24,PLC TO FOLLOW RAMP Breakpoints A to B
        [30].3   // FV24,Current vessel deferred chilling active
        [19]   // FV24,Current FV max. fermentation time
        [41]   // FV24,Cone ACTUAL TEMPERATURE -DEGREES 'C'*10
        [20]   // FV24,Current FV warm conditioning time
        [28]   // FV24,CURRENT VOLUME HL*10
        [15].3   // FV24,PLC TO USE CONE COOLING JACKET
        [30].1   // FV24,Cone Cooling Valve to open
        [26]   // FV24,Calculated Setpoint 1/10 degrees C
        [10]   // FV24,TEMPERATURE SETPOINT E. 1/10 DEGREE 'C'
        [12]   // FV24,TEMPERATURE SETPOINT F. 1/10 DEGREE 'C'
        [14]   // FV24,TEMPERATURE SETPOINT G. 1/10 DEGREE 'C'
        [30].0   // FV24,Jacket Cooling Valve to open
        [24]   // FV24,Phase0=No control 1to6 =Fermenting 8 =Pitching Hold 10 =Maturation 11to16=Conditioning
        [0]   // FV24,FV SYSTEM WORKING BUFFER VESSEL NUMBER
        [2]   // FV24,TEMPERATURE SETPOINT A. 1/10 DEGREE 'C'
        [30].4   // FV24,Current vessel final temp.reached
        [4]   // FV24,TEMPERATURE SETPOINT B. 1/10 DEGREE 'C'
        [36]   // FV24,Current vessel time to deferred chlling start (hrs.x10)
        [6]   // FV24,TEMPERATURE SETPOINT C. 1/10 DEGREE 'C'
        [8]   // FV24,TEMPERATURE SETPOINT D. 1/10 DEGREE 'C'
        [29]   // FV24,FLAGS - PLC CONTROL
        [27]   // FV24,CURRENT ELAPSED HOURS *10
        [22]   // FV24,Current FV total residence time
        [40]   // FV24,FV Routing Status 9=Dirty
        [29].0   // FV24,PC TO SAVE TEMPERATURE DATA
        [16].1   // FV24,Profile control flag Hold at B.P B
        [16].2   // FV24,Profile control flag Hold at B.P C
        [16].3   // FV24,Profile control flag Hold at B.P D
        [16].4   // FV24,Profile control flag Hold at B.P E
        [16].5   // FV24,Profile control flag Hold at B.P F
        [16].6   // FV24,Profile control flag Hold at B.P G
        [11]   // FV24,TEMPERATURE BREAKPOINT F. TIME 1/10 HOURS(ALWAYS=0)
        [13]   // FV24,TEMPERATURE BREAKPOINT G. TIME 1/10 HOURS(ALWAYS=0)
        [30].5   // FV24,Current vessel deferred chilling temp.high flag
        [15].9   // FV24,Current vessel deferred chilling manual override
        [1]   // FV24,TEMPERATURE BREAKPOINT A. TIME 1/10 HOURS(ALWAYS=0)
        [29].1   // FV24,Current vessel deferred chilling enabled flag
        [3]   // FV24,TEMPERATURE BREAKPOINT B. TIME 1/10 HOURS(ALWAYS=0)
        [5]   // FV24,TEMPERATURE BREAKPOINT C. TIME 1/10 HOURS(ALWAYS=0)
        [7]   // FV24,TEMPERATURE BREAKPOINT D. TIME 1/10 HOURS(ALWAYS=0)
        [9]   // FV24,TEMPERATURE BREAKPOINT E. TIME 1/10 HOURS(ALWAYS=0)
   FV_N135 : INT[50] := ([0] := 25, [1] := -32767, [2] := -32767, [3] := -32767, [4] := -32767, [5] := -32767, [6] := -32767, [7] := -32767, [8] := -32767, [9] := -32767, [10] := -32767, [11] := -32767, [12] := -32767, [13] := -32767, [14] := -32767, [15] := -32767, [16] := -32767, [17] := -32767, [18] := -32767, [19] := -32767, [20] := -32767, [21] := -32767, [22] := -32767, [23] := 2, [25] := 222, [30] := 32);   // FV25, CURRENT FV DATA
        [15]   // FV25,FLAGS-PROFILE CONTROL
        [15].4   // FV25,Profile Control Flags : This is a maturation profile
        [15].5   // FV25,Profile Control Flags : This is a conditioning profile
        [25]   // FV25,Jacket ACTUAL TEMPERATURE -DEGREES 'C'*10
        [15].2   // FV25,PLC TO FOLLOW RAMP Breakpoints A to B
        [19]   // FV25,Current FV max. fermentation time
        [30].3   // FV25,Current vessel deferred chilling active
        [20]   // FV25,Current FV warm conditioning time
        [41]   // FV25,Cone ACTUAL TEMPERATURE -DEGREES 'C'*10
        [15].3   // FV25,PLC TO USE CONE COOLING JACKET
        [28]   // FV25,CURRENT VOLUME HL*10
        [26]   // FV25,Calculated Setpoint 1/10 degrees C
        [30].1   // FV25,Cone Cooling Valve to open
        [10]   // FV25,TEMPERATURE SETPOINT E. 1/10 DEGREE 'C'
        [12]   // FV25,TEMPERATURE SETPOINT F. 1/10 DEGREE 'C'
        [14]   // FV25,TEMPERATURE SETPOINT G. 1/10 DEGREE 'C'
        [24]   // FV25,Phase0=No control 1to6 =Fermenting 8 =Pitching Hold 10 =Maturation 11to16=Conditioning
        [30].0   // FV25,Jacket Cooling Valve to open
        [0]   // FV25,FV SYSTEM WORKING BUFFER VESSEL NUMBER
        [2]   // FV25,TEMPERATURE SETPOINT A. 1/10 DEGREE 'C'
        [30].4   // FV25,Current vessel final temp.reached
        [4]   // FV25,TEMPERATURE SETPOINT B. 1/10 DEGREE 'C'
        [6]   // FV25,TEMPERATURE SETPOINT C. 1/10 DEGREE 'C'
        [8]   // FV25,TEMPERATURE SETPOINT D. 1/10 DEGREE 'C'
        [36]   // FV25,Current vessel time to deferred chlling start (hrs.x10)
        [27]   // FV25,CURRENT ELAPSED HOURS *10
        [40]   // FV25,FV Routing Status 9=Dirty
        [29]   // FV25,FLAGS - PLC CONTROL
        [22]   // FV25,Current FV total residence time
        [16].1   // FV25,Profile control flag Hold at B.P B
        [16].2   // FV25,Profile control flag Hold at B.P C
        [16].3   // FV25,Profile control flag Hold at B.P D
        [16].4   // FV25,Profile control flag Hold at B.P E
        [29].0   // FV25,PC TO SAVE TEMPERATURE DATA
        [16].5   // FV25,Profile control flag Hold at B.P F
        [16].6   // FV25,Profile control flag Hold at B.P G
        [11]   // FV25,TEMPERATURE BREAKPOINT F. TIME 1/10 HOURS(ALWAYS=0)
        [13]   // FV25,TEMPERATURE BREAKPOINT G. TIME 1/10 HOURS(ALWAYS=0)
        [30].5   // FV25,Current vessel deferred chilling temp.high flag
        [1]   // FV25,TEMPERATURE BREAKPOINT A. TIME 1/10 HOURS(ALWAYS=0)
        [29].1   // FV25,Current vessel deferred chilling enabled flag
        [3]   // FV25,TEMPERATURE BREAKPOINT B. TIME 1/10 HOURS(ALWAYS=0)
        [5]   // FV25,TEMPERATURE BREAKPOINT C. TIME 1/10 HOURS(ALWAYS=0)
        [7]   // FV25,TEMPERATURE BREAKPOINT D. TIME 1/10 HOURS(ALWAYS=0)
        [15].9   // FV25,Current vessel deferred chilling manual override
        [9]   // FV25,TEMPERATURE BREAKPOINT E. TIME 1/10 HOURS(ALWAYS=0)
   FV_N136 : INT[50] := ([0] := 26, [2] := 30, [3] := 240, [4] := 30, [5] := 480, [6] := 30, [7] := 720, [8] := 30, [9] := 960, [10] := 30, [11] := 1200, [12] := 30, [13] := 32767, [14] := 30, [15] := 20, [17] := -32767, [18] := -32767, [20] := 1492, [22] := 1492, [23] := 1, [24] := 10, [25] := 46, [26] := 30, [27] := 1492, [30] := 57);   // YSV1, CURRENT FV DATA
        [15]   // YSV1,FLAGS-PROFILE CONTROL
        [15].4   // YSV1,Profile Control Flags : This is a maturation profile
        [25]   // YSV1,Jacket ACTUAL TEMPERATURE -DEGREES 'C'*10
        [15].5   // YSV1,Profile Control Flags : This is a conditioning profile
        [15].2   // YSV1,PLC TO FOLLOW RAMP Breakpoints A to B
        [19]   // YSV1,Current FV max. fermentation time
        [30].3   // YSV1,Current vessel deferred chilling active
        [20]   // YSV1,Current FV warm conditioning time
        [41]   // YSV1,Cone ACTUAL TEMPERATURE -DEGREES 'C'*10
        [15].3   // YSV1,PLC TO USE CONE COOLING JACKET
        [26]   // YSV1,Calculated Setpoint 1/10 degrees C
        [28]   // YSV1,CURRENT VOLUME HL*10
        [10]   // YSV1,TEMPERATURE SETPOINT E. 1/10 DEGREE 'C'
        [12]   // YSV1,TEMPERATURE SETPOINT F. 1/10 DEGREE 'C'
        [30].1   // YSV1,Cone Cooling Valve to open
        [14]   // YSV1,TEMPERATURE SETPOINT G. 1/10 DEGREE 'C'
        [24]   // YSV1,Phase0=No control 1to6 =Fermenting 8 =Pitching Hold 10 =Maturation 11to16=Conditioning
        [0]   // YSV1,FV SYSTEM WORKING BUFFER VESSEL NUMBER
        [2]   // YSV1,TEMPERATURE SETPOINT A. 1/10 DEGREE 'C'
        [30].4   // YSV1,Current vessel final temp.reached
        [4]   // YSV1,TEMPERATURE SETPOINT B. 1/10 DEGREE 'C'
        [6]   // YSV1,TEMPERATURE SETPOINT C. 1/10 DEGREE 'C'
        [30].0   // YSV1,Jacket Cooling Valve to open
        [8]   // YSV1,TEMPERATURE SETPOINT D. 1/10 DEGREE 'C'
        [36]   // YSV1,Current vessel time to deferred chlling start (hrs.x10)
        [27]   // YSV1,CURRENT ELAPSED HOURS *10
        [40]   // YSV1,FV Routing Status 9=Dirty
        [29]   // YSV1,FLAGS - PLC CONTROL
        [22]   // YSV1,Current FV total residence time
        [29].0   // YSV1,PC TO SAVE TEMPERATURE DATA
        [16].1   // YSV1,Profile control flag Hold at B.P B
        [16].2   // YSV1,Profile control flag Hold at B.P C
        [16].3   // YSV1,Profile control flag Hold at B.P D
        [16].4   // YSV1,Profile control flag Hold at B.P E
        [16].5   // YSV1,Profile control flag Hold at B.P F
        [16].6   // YSV1,Profile control flag Hold at B.P G
        [1]   // YSV1,TEMPERATURE BREAKPOINT A. TIME 1/10 HOURS(ALWAYS=0)
        [11]   // YSV1,TEMPERATURE BREAKPOINT F. TIME 1/10 HOURS(ALWAYS=0)
        [13]   // YSV1,TEMPERATURE BREAKPOINT G. TIME 1/10 HOURS(ALWAYS=0)
        [30].5   // YSV1,Current vessel deferred chilling temp.high flag
        [29].1   // YSV1,Current vessel deferred chilling enabled flag
        [3]   // YSV1,TEMPERATURE BREAKPOINT B. TIME 1/10 HOURS(ALWAYS=0)
        [5]   // YSV1,TEMPERATURE BREAKPOINT C. TIME 1/10 HOURS(ALWAYS=0)
        [7]   // YSV1,TEMPERATURE BREAKPOINT D. TIME 1/10 HOURS(ALWAYS=0)
        [9]   // YSV1,TEMPERATURE BREAKPOINT E. TIME 1/10 HOURS(ALWAYS=0)
        [15].9   // YSV1,Current vessel deferred chilling manual override
   FV_N137 : INT[50] := ([0] := 27, [2] := 30, [3] := 240, [4] := 30, [5] := 480, [6] := 30, [7] := 720, [8] := 30, [9] := 960, [10] := 30, [11] := 1200, [12] := 30, [13] := 32767, [14] := 30, [15] := 20, [17] := -32767, [18] := -32767, [20] := 303, [22] := 303, [23] := 1, [24] := 10, [25] := 31, [26] := 30, [27] := 303, [30] := 25);   // YSV2, CURRENT FV DATA
        [15]   // YSV2,FLAGS-PROFILE CONTROL
        [15].4   // YSV2,Profile Control Flags : This is a maturation profile
        [25]   // YSV2,Jacket ACTUAL TEMPERATURE -DEGREES 'C'*10
        [15].5   // YSV2,Profile Control Flags : This is a conditioning profile
        [15].2   // YSV2,PLC TO FOLLOW RAMP Breakpoints A to B
        [19]   // YSV2,Current FV max. fermentation time
        [20]   // YSV2,Current FV warm conditioning time
        [30].3   // YSV2,Current vessel deferred chilling active
        [41]   // YSV2,Cone ACTUAL TEMPERATURE -DEGREES 'C'*10
        [10]   // YSV2,TEMPERATURE SETPOINT E. 1/10 DEGREE 'C'
        [15].3   // YSV2,PLC TO USE CONE COOLING JACKET
        [26]   // YSV2,Calculated Setpoint 1/10 degrees C
        [28]   // YSV2,CURRENT VOLUME HL*10
        [12]   // YSV2,TEMPERATURE SETPOINT F. 1/10 DEGREE 'C'
        [14]   // YSV2,TEMPERATURE SETPOINT G. 1/10 DEGREE 'C'
        [30].0   // YSV2,Jacket Cooling Valve to open
        [30].1   // YSV2,Cone Cooling Valve to open
        [24]   // YSV2,Phase0=No control 1to6 =Fermenting 8 =Pitching Hold 10 =Maturation 11to16=Conditioning